                                   //current limit or reason for switch off output 6
                                   IF #statHMI.stateOutput6 = #CONST_STATE_OUT_AUTO_SWITCHED_OFF OR
                                       #statHMI.stateOutput6 = #CONST_STATE_OUT_RESET_POSSIBLE
                                   THEN
                                       #statHMI.reasonOutputSwitchedOff6 := BYTE_TO_INT(#statOutputCurrentLimit6);
                                   ELSE
                                       #statHMI.outputCurrentLimit6 := (BYTE_TO_INT(#statOutputCurrentLimit6) * #statHMI.nominalOutputCurrent) / #CONST_CONVERT_CURRENT;
                                   END_IF;

                                   //current limit or reason for switch off output 7
                                   IF #statHMI.stateOutput7 = #CONST_STATE_OUT_AUTO_SWITCHED_OFF OR
                                       #statHMI.stateOutput7 = #CONST_STATE_OUT_RESET_POSSIBLE
                                   THEN
                                       #statHMI.reasonOutputSwitchedOff7 := BYTE_TO_INT(#statOutputCurrentLimit7);
                                   ELSE
                                       #statHMI.outputCurrentLimit7 := (BYTE_TO_INT(#statOutputCurrentLimit7) * #statHMI.nominalOutputCurrent) / #CONST_CONVERT_CURRENT;
                                   END_IF;

                                   //current limit or reason for switch off output 8
                                   IF #statHMI.stateOutput8 = #CONST_STATE_OUT_AUTO_SWITCHED_OFF OR
                                       #statHMI.stateOutput8 = #CONST_STATE_OUT_RESET_POSSIBLE
                                   THEN
                                       #statHMI.reasonOutputSwitchedOff8 := BYTE_TO_INT(#statOutputCurrentLimit8);
                                   ELSE
                                       #statHMI.outputCurrentLimit8 := (BYTE_TO_INT(#statOutputCurrentLimit8) * #statHMI.nominalOutputCurrent) / #CONST_CONVERT_CURRENT;
                                   END_IF;

                               END_IF;

                           ELSE
                               // wrong frame Id
                               #statErrorFrameID := true;
                           END_IF;

                           IF #statGetFrame.frame0 = TRUE
                               AND #statGetFrame.frame1 = TRUE
                               AND #statGetFrame.frame2 = TRUE
                               AND #statGetFrame.frame3 = TRUE
                           THEN

                               #statIndexArticleNumber := 1;

                               FOR #statIndexArticleNumber := #CONST_START_CNT_INDEX1 TO #CONST_END_CNT_INDEX18 BY 1 DO
                                   IF #statArticleNumber[#statIndexArticleNumber] <> #statArticleNumberOld[#statIndexArticleNumber]
                                   THEN
                                       #statNewArticleNumberDetected := true;
                                   END_IF;
                               END_FOR;


                               IF #statNewArticleNumberDetected = TRUE
                               THEN

                                   #statNewArticleNumberDetected := false;
                                   #statArticleNumberChanged := true;

                                   Chars_TO_Strg(Chars := #statArticleNumber,
                                                 pChars := 0,
                                                 Cnt := 0,
                                                 Strg => #statHMI.articleNumber);
                                   #statArticleNumberOld := #statArticleNumber;
                               END_IF;


                               IF #statFabricationPlace = TRUE
                               THEN
                                   //fabrication place: Sibiu
                                   #statSerialNumber[1] := 'Y';
                                   #statSerialNumber[2] := 'S';
                                   #statSerialNumber[3] := 'U';
                                   #statSerialNumber[4] := '/';
                                   #statSerialNumber[5] := #statConstructionYearChar;
                                   #statSerialNumber[6] := #statConstructionMonthChar;
                                   #statSerialNumber[7] := ' ';
                                   #statSerialNumber[8] := ' ';
                                   #statSerialNumber[9] := ' ';
                                   #statSerialNumber[10] := ' ';
                                   #statSerialNumber[11] := ' ';
                                   #statSerialNumber[12] := ' ';
                                   #statSerialNumber[13] := ' ';
                               ELSE
                                   //fabrication place: Vienna
                                   #statSerialNumber[1] := 'Q';
                                   #statSerialNumber[2] := '6';
                                   #statSerialNumber[3] := '/';
                                   #statSerialNumber[4] := #statConstructionYearChar;
                                   #statSerialNumber[5] := #statConstructionMonthChar;
                                   #statSerialNumber[6] := ' ';
                                   #statSerialNumber[7] := ' ';
                                   #statSerialNumber[8] := ' ';
                                   #statSerialNumber[9] := ' ';
                                   #statSerialNumber[10] := ' ';
                                   #statSerialNumber[11] := ' ';
                                   #statSerialNumber[12] := ' ';
                                   #statSerialNumber[13] := ' ';

                               END_IF;

                               #statIndexSerialNumber := 1;

                               FOR #statIndexSerialNumber := #CONST_START_CNT_INDEX1 TO #CONST_END_CNT_INDEX13 BY 1 DO
                                   IF #statSerialNumber[#statIndexSerialNumber] <> #statSerialNumberOld[#statIndexSerialNumber]
                                   THEN
                                       #statNewSerialNumberDetected := true;
                                   END_IF;
                               END_FOR;

                               IF #statNewSerialNumberDetected = TRUE
                               THEN
                                   #statNewSerialNumberDetected := false;
                                   Chars_TO_Strg(Chars := #statSerialNumber,
                                                 pChars := 0,
                                                 Cnt := 0,
                                                 Strg => #statHMI.serialNumber);
                                   #statSerialNumberOld := #statSerialNumber;
                               END_IF;

                               #statGetFrame.frame0 := FALSE;
                               #statGetFrame.frame1 := FALSE;
                               #statGetFrame.frame2 := FALSE;
                               #statGetFrame.frame3 := FALSE;
                           END_IF;

                           // set output data structure
                           #HMI.deviceName := #statHMI.deviceName;
                           #HMI.stateCOM := true;
                           #HMI.stateDipSwitchTD1 := #statHMI.stateDipSwitchTD1;
                           #HMI.stateDipSwitchTD2 := #statHMI.stateDipSwitchTD2;
                           #HMI.stateOutput1 := #statHMI.stateOutput1;
                           #HMI.stateOutput2 := #statHMI.stateOutput2;
                           #HMI.stateOutput3 := #statHMI.stateOutput3;
                           #HMI.stateOutput4 := #statHMI.stateOutput4;
                           #HMI.stateOutput5 := #statHMI.stateOutput5;
                           #HMI.stateOutput6 := #statHMI.stateOutput6;
                           #HMI.stateOutput7 := #statHMI.stateOutput7;
                           #HMI.stateOutput8 := #statHMI.stateOutput8;
                           #HMI.outputCurrent1 := #statHMI.outputCurrent1;
                           #HMI.outputCurrent2 := #statHMI.outputCurrent2;
                           #HMI.outputCurrent3 := #statHMI.outputCurrent3;
                           #HMI.outputCurrent4 := #statHMI.outputCurrent4;
                           #HMI.outputCurrent5 := #statHMI.outputCurrent5;
                           #HMI.outputCurrent6 := #statHMI.outputCurrent6;
                           #HMI.outputCurrent7 := #statHMI.outputCurrent7;
                           #HMI.outputCurrent8 := #statHMI.outputCurrent8;
                           #HMI.outputCurrentLimit1 := #statHMI.outputCurrentLimit1;
                           #HMI.outputCurrentLimit2 := #statHMI.outputCurrentLimit2;
                           #HMI.outputCurrentLimit3 := #statHMI.outputCurrentLimit3;
                           #HMI.outputCurrentLimit4 := #statHMI.outputCurrentLimit4;
                           #HMI.outputCurrentLimit5 := #statHMI.outputCurrentLimit5;
                           #HMI.outputCurrentLimit6 := #statHMI.outputCurrentLimit6;
                           #HMI.outputCurrentLimit7 := #statHMI.outputCurrentLimit7;
                           #HMI.outputCurrentLimit8 := #statHMI.outputCurrentLimit8;
                           #HMI.reasonOutputSwitchedOff1 := #statHMI.reasonOutputSwitchedOff1;
                           #HMI.reasonOutputSwitchedOff2 := #statHMI.reasonOutputSwitchedOff2;
                           #HMI.reasonOutputSwitchedOff3 := #statHMI.reasonOutputSwitchedOff3;
                           #HMI.reasonOutputSwitchedOff4 := #statHMI.reasonOutputSwitchedOff4;
                           #HMI.reasonOutputSwitchedOff5 := #statHMI.reasonOutputSwitchedOff5;
                           #HMI.reasonOutputSwitchedOff6 := #statHMI.reasonOutputSwitchedOff6;
                           #HMI.reasonOutputSwitchedOff7 := #statHMI.reasonOutputSwitchedOff7;
                           #HMI.reasonOutputSwitchedOff8 := #statHMI.reasonOutputSwitchedOff8;
                           #HMI.nominalOutputCurrent := #statHMI.nominalOutputCurrent;
                           #HMI.productState := #statHMI.productState;
                           #HMI.firmwareVersion := #statHMI.firmwareVersion;
                           #HMI.startup := #statHMI.startup;
                           #HMI.outputNumber := #statHMI.outputNumber;
                           #HMI.stateReset := #statHMI.stateReset;
                           #HMI.articleNumber := #statHMI.articleNumber;
                           #HMI.serialNumber := #statHMI.serialNumber;

                       ELSE
                           //wrong device (no PSU OR SEL)
                           #statErrorDevice := true;
                       END_IF;
                       #statFrameOld := #statFrame;
                   END_IF;

               ELSE

                   IF #statInit = true
                   THEN
                       #statErrorFrameLength := true;
                   END_IF;

               END_IF;


               #statArrayImpulse[0] := #statTimeSave.deltaTimeImpulse;

               FOR #statIndexResetImpulse := #CONST_START_CNT_INDEX1 TO #CONST_END_CNT_INDEX63 BY 1 DO
                   #statArrayImpulse[#statIndexResetImpulse] := #CONST_TIME_0;
               END_FOR;

               FOR #statIndexResetPause := #CONST_START_CNT_INDEX0 TO #CONST_END_CNT_INDEX63 BY 1 DO
                   #statArrayPause[#statIndexResetPause] := #CONST_TIME_0;
               END_FOR;

               #statStartTimerWait := true;
               #statNoEvaluation := true;

               //Impulse detection    
           ELSIF #statTimeSave.deltaTimeImpulse >= #CONST_IMPULSE_MIN
               AND #statTimeSave.deltaTimeImpulse <= #CONST_IMPULSE_MAX
               AND #statImpulseDetected = TRUE
           THEN
               #statImpulseDetected := false;
               #statIndexResetImpulse := #CONST_INT_1;

               //save time of impulses to check frame length
               #statArrayImpulse[#statIndexImpulse] := #statTimeSave.deltaTimeImpulse;
               #statIndexImpulse := #statIndexImpulse + #CONST_INT_1;

               //count number of impulses
               #statCntImpulse := #statCntImpulse + #CONST_INT_1;

           END_IF;


           IF #statPauseDetected = TRUE
           THEN
               #statPauseDetected := false;
               #statIndexResetPause := #CONST_INT_0;

               //save time of pauses to check frame length
               #statArrayPause[#statIndexPause] := #statTimeSave.deltaTimePause;
               #statIndexPause := #statIndexPause + #CONST_INT_1;

               //count number of pauses
               #statCntPause := #statCntPause + #CONST_INT_1;

           END_IF;

           // bit detection
           IF #statNoEvaluation = false
               AND #statFrameEvaluationStopp = false
               AND ((#statPosEdgeDetectedTrigger = true)
               OR (#statNegEdgeDetectedTrigger = true))
           THEN

               IF #statPosEdgeDetectedTrigger = true
               THEN
                   #statArrayBits[#statCntBits] := true;
               ELSIF #statNegEdgeDetectedTrigger = true
               THEN
                   #statArrayBits[#statCntBits] := false;
               END_IF;

               #statStartTimerWait := true;
               #statNoEvaluation := true;

               IF (#statCntBits >= (#CONST_CNT_BITS_MAX - #CONST_INT_1))
               THEN
                   #statFrameEvaluationStopp := true;
                   #statCntBits := #CONST_INT_0;
               ELSE
                   #statCntBits := #statCntBits + #CONST_INT_1;
               END_IF;

           END_IF;

           //check max number of impulses and pauses in frame
           IF #statCntImpulse > #CONST_CNT_BITS_MAX
           THEN
               #statIndexImpulse := #CONST_INT_1;
               #statErrorFrameContent := TRUE;
           END_IF;

           IF #statCntPause > #CONST_CNT_PAUSE_MAX
           THEN
               #statIndexPause := #CONST_INT_0;
               #statErrorFrameContent := true;
           END_IF;

           IF #statErrorFrameContent = TRUE
           THEN
               #statStatusInt := #CONST_ERR_FRAMECONTENT;
               #statErrorInt := true;
           ELSIF #statErrorFrameLength = TRUE
           THEN
               #statStatusInt := #CONST_ERR_FRAMELENGTH;
               #statErrorInt := true;
           ELSIF #statErrorDevice = TRUE
           THEN
               #statStatusInt := #CONST_ERR_DEVICE;
               #statErrorInt := true;
           ELSIF #statErrorFrameID = TRUE
           THEN
               #statStatusInt := #CONST_ERR_FRAME_ID;
               #statErrorInt := true;
           ELSIF #statArticleNumberChanged = TRUE
           THEN
               #statStatusInt := #CONST_ERR_ARTICLE_NUMBER;
               #statErrorInt := true;
           END_IF;

           IF #statErrorInt = TRUE
           THEN
               #statErrorFrameLength := false;
               #statErrorFrameContent := false;
               #statErrorDevice := false;
               #statErrorFrameID := FALSE;
               #statArticleNumberChanged := false;
               #statStateIndex := #STATE_ERROR;
           END_IF;

       #STATE_ERROR:
           #statError := true;
           #statBusy := false;
           #statDone := false;
           #statStatus := #statStatusInt;
           #statStatusInt := #CONST_WORD_0;
           #statStartTimerSys := false;
           #statIndexResetBitArray := #CONST_INT_0;
           #statStartWatchDogTimerNeg := false;
           #statStartWatchDogTimerPos := false;

           IF #statErrorInt = TRUE
           THEN
               #statStateIndex := #STATE_EVALUATION;
               #statErrorInt := false;
               #statStartWatchDogTimerNeg := true;
               #statStartWatchDogTimerPos := true;
           ELSE
               #statStateIndex := #STATE_IDLE;
           END_IF;

       ELSE  // Statement section ELSE
           #statIndexResetBitArray := #CONST_INT_0;
           #statStateIndex := #STATE_IDLE;
   END_CASE;


   //Timer
   #instTimerWait(IN := #statStartTimerWait,
                  PT := #CONST_TIME_WAIT);

   IF #instTimerWait.Q = TRUE
   THEN
       #statStartTimerWait := false;
       #statNoEvaluation := false;
   END_IF;

   #instSysTimer(IN := #statStartTimerSys,
                 PT := #CONST_SYS_TIMER);


   IF #instSysTimer.Q = TRUE
   THEN
       #statStatusInt := #CONST_ERR_CYCLE_TIME;
       #statStateIndex := #STATE_ERROR;
   END_IF;

   #instWatchDogTimerPos(IN := #statStartWatchDogTimerPos,
                         PT := #CONST_WATCHDOG_TIMER);

   #instWatchDogTimerNeg(IN := #statStartWatchDogTimerNeg,
                         PT := #CONST_WATCHDOG_TIMER);

   IF #instWatchDogTimerNeg.Q = TRUE
       OR #instWatchDogTimerPos.Q = TRUE
   THEN
       #statStatusInt := #CONST_ERR_WATCHDOG;
       #statStateIndex := #STATE_ERROR;

       IF #HMI.stateNoCommunication = FALSE
       THEN
           #HMI.stateNoCommunication := true;

           #HMI.deviceName := #CONST_DEVICE_NAME_DEFAULT;
           #HMI.stateCOM := true;
           #HMI.stateDipSwitchTD1 := FALSE;
           #HMI.stateDipSwitchTD2 := FALSE;
           #HMI.stateOutput1 := #CONST_STATE_OUT_DEFAULT;
           #HMI.stateOutput2 := #CONST_STATE_OUT_DEFAULT;
           #HMI.stateOutput3 := #CONST_STATE_OUT_DEFAULT;
           #HMI.stateOutput4 := #CONST_STATE_OUT_DEFAULT;
           #HMI.stateOutput5 := #CONST_STATE_OUT_DEFAULT;
           #HMI.stateOutput6 := #CONST_STATE_OUT_DEFAULT;
           #HMI.stateOutput7 := #CONST_STATE_OUT_DEFAULT;
           #HMI.stateOutput8 := #CONST_STATE_OUT_DEFAULT;
           #HMI.outputCurrent1 := #CONST_CURRENT_OUT_DEFAULT;
           #HMI.outputCurrent2 := #CONST_CURRENT_OUT_DEFAULT;
           #HMI.outputCurrent3 := #CONST_CURRENT_OUT_DEFAULT;
           #HMI.outputCurrent4 := #CONST_CURRENT_OUT_DEFAULT;
           #HMI.outputCurrent5 := #CONST_CURRENT_OUT_DEFAULT;
           #HMI.outputCurrent6 := #CONST_CURRENT_OUT_DEFAULT;
           #HMI.outputCurrent7 := #CONST_CURRENT_OUT_DEFAULT;
           #HMI.outputCurrent8 := #CONST_CURRENT_OUT_DEFAULT;
           #HMI.outputCurrentLimit1 := #CONST_CURRENT_OUT_DEFAULT;
           #HMI.outputCurrentLimit2 := #CONST_CURRENT_OUT_DEFAULT;
           #HMI.outputCurrentLimit3 := #CONST_CURRENT_OUT_DEFAULT;
           #HMI.outputCurrentLimit4 := #CONST_CURRENT_OUT_DEFAULT;
           #HMI.outputCurrentLimit5 := #CONST_CURRENT_OUT_DEFAULT;
           #HMI.outputCurrentLimit6 := #CONST_CURRENT_OUT_DEFAULT;
           #HMI.outputCurrentLimit7 := #CONST_CURRENT_OUT_DEFAULT;
           #HMI.outputCurrentLimit8 := #CONST_CURRENT_OUT_DEFAULT;
           #HMI.reasonOutputSwitchedOff1 := #CONST_REASON_SWITCHED_OFF_DEFAULT;
           #HMI.reasonOutputSwitchedOff2 := #CONST_REASON_SWITCHED_OFF_DEFAULT;
           #HMI.reasonOutputSwitchedOff3 := #CONST_REASON_SWITCHED_OFF_DEFAULT;
           #HMI.reasonOutputSwitchedOff4 := #CONST_REASON_SWITCHED_OFF_DEFAULT;
           #HMI.reasonOutputSwitchedOff5 := #CONST_REASON_SWITCHED_OFF_DEFAULT;
           #HMI.reasonOutputSwitchedOff6 := #CONST_REASON_SWITCHED_OFF_DEFAULT;
           #HMI.reasonOutputSwitchedOff7 := #CONST_REASON_SWITCHED_OFF_DEFAULT;
           #HMI.reasonOutputSwitchedOff8 := #CONST_REASON_SWITCHED_OFF_DEFAULT;
           #HMI.nominalOutputCurrent := #CONST_NOMINAL_CURRENT3;
           #HMI.productState := #CONST_FW_PRODUCT_STATE_DEFAULT;
           #HMI.firmwareVersion := #CONST_FW_PRODUCT_STATE_DEFAULT;
           #HMI.startup := #CONST_STARTUP_DEFAULT;
           #HMI.outputNumber := #CONST_OUTPUT_NUMBER_4;
           #HMI.stateReset := FALSE;
           #HMI.articleNumber := #CONST_ARTICLE_NUMBER_DEFAULT;
           #HMI.serialNumber := #CONST_SERIAL_NUMBER_DEFAULT;

       END_IF;

   END_IF;

   #instTimerReset(IN:=#reset,
                   PT:=#CONST_RESET_TIMER);


   //edge Control
   #statImpulseOld := #impulse;
   #statPosEdgeDetectedTrigger := false;
   #statNegEdgeDetectedTrigger := false;

   //Cycle Time Control
   #statTimeSave.sysTimeOld := #statTimeSave.sysTime;

   // set outputs
   IF #HMI.setReset = TRUE
   THEN
       #HMI.setReset := false;
       #reset := true;
   ELSE
       IF #instTimerReset.Q = TRUE
       THEN
           #reset := false;
       END_IF;
   END_IF;

   #busy := #statBusy;
   #error := #statError;
   #done := #statDone;
   #status := #statStatus;
END_REGION
END_FUNCTION_BLOCK

FUNCTION_BLOCK "LPSE"   // FB6970, LAD
{ S7_Optimized_Access := 'TRUE' }
VERSION : 0.1
   VAR_INPUT
      impulse : Bool;
      reset : Bool;
   END_VAR
   VAR_OUTPUT
      done : Bool;
      busy : Bool;
      status : Word;
      error : Bool;
   END_VAR
   VAR
      statImpulseOld : Bool;
      HMI : Struct
         channelstate : Byte;
      END_STRUCT;
      statResetOld : Bool;
      statTimeSaver : Struct
         TimeTckRisingEdge : DTL;
         TimeTckFallingEdge : DTL;
         RisingEdgeDetected : Bool;
         FallingEdgeDetected : Bool;
         stateEdge : Int := 0;
      END_STRUCT;
      statDeltaTimeImpulse : Time;
      statDeltaTimePause : Time;
      statStartImpulseDetected : Bool;
      statImpulseDetected : Bool;
      statChannelState : Byte;
      statTimePauseSave0 : Time;
      statTimePauseSave1 : Time;
      statTimePauseSave2 : Time;
      statTimePauseSave3 : Time;
      statTimePauseSave4 : Time;
      statTimeImpulseSave0 : Time;
      statTimeImpulseSave1 : Time;
      statTimeImpulseSave2 : Time;
      statTimeImpulseSave3 : Time;
      statTimeImpulseSave4 : Time;
      statFrameImulseDetected : Bool;
      statNumberOfImpulses : Int;
      statChannelActive1 : Bool;
      statChannelActive2 : Bool;
      statChannelActive3 : Bool;
      statChannelActive4 : Bool;
      statCountChannelPos : Int;
      statCurrentPos1 : Int;
      statCurrentPos2 : Int;
      statCurrentPos3 : Int;
      statCurrentPos4 : Int;
      statTimeToImpulse : Time;
      statTimePause : Time;
      statTimeImpulse : Time;
      statTimeFrame : Time;
      statFrameOk : Bool;
      statCycleTimeNok : Bool;
      statDeltaSysTime : Time;
      instSysTimer : TON_TIME;
      statSysTimerStart : Bool;
      statSysTimerStop : Bool;
      statStatus : Word;
      statIndex : Int;
      statSysTimerRun : Time;
      instWatchDogTimerRising : TON_TIME;
      statWatchDogTimerRisingStart : Bool;
      statWatchDogTimerRisingStop : Bool;
      statWatchDogTimerRisingRun : Time;
      statResetRequest : Bool;
      statSysTimeDtl : DTL;
      statSysTimeOldDtl : DTL;
      instWatchDogTimerFalling : TON_TIME;
      statWatchDogTimerFallingStart : Bool;
      statWatchDogTimerFallingStop : Bool;
      statWatchDogTimerFallingRun : Time;
   END_VAR
   VAR_TEMP
      tempRetvalRdSys : Int;
      tempRetvalRdSysPosEdge : Int;
      tempRetvalRdSysNegEdge : Int;
      tempLatchTime : DTL;
      tempSysTime : DTL;
   END_VAR
   VAR CONSTANT
      STATE_IDLE : Int := 0;
      STATE_EVALUATION : Int := 1;
      STATE_ERROR : Int := 2;
      TIME_FRAME_MAX : Time := T#2850ms;
      TIME_FRAME_MIN : Time := T#2650ms;
      TIME_STARTIMPULSE_MIN : Time := T#400ms;
      TIME_STARTIMPULSE_MAX : Time := T#600ms;
      TIME_IMPULSE_MIN : Time := T#150ms;
      TIME_IMPULSE_MAX : Time := T#350ms;
      TIME_PAUSE1_MIN : Time := T#150ms;
      TIME_PAUSE1_MAX : Time := T#350ms;
      TIME_PAUSE2_MIN : Time := T#650ms;
      TIME_PAUSE2_MAX : Time := T#850ms;
      TIME_PAUSE3_MIN : Time := T#1150ms;
      TIME_PAUSE3_MAX : Time := T#1350ms;
      TIME_PAUSE4_MIN : Time := T#1650ms;
      TIME_PAUSE4_MAX : Time := T#1850ms;
      TIME_PAUSE_FRAME_MAX : Time := T#2350ms;
      TIME_PAUSE_FRAME_MIN : Time := T#2150ms;
      CONST_TIME_102 : Time := T#102ms;
      CONST_TIME_0 : Time := t#0ms;
      CONST_STATE_RISING_EDGE : Int := 15;
      CONST_STATE_FALLING_EDGE : Int := 16;
      CONST_WORD_0 : Word := 16#0000;
      CONST_BYTE_0 : Byte := 16#00;
      CONST_INT_0 : Int := 0;
      CONST_CHANNEL_POS4 : Int := 4;
      CONST_CHANNEL_POS1 : Int := 1;
      CONST_CHANNEL_POS2 : Int := 2;
      CONST_CHANNEL_POS3 : Int := 3;
      CONST_WATCHDOG_TIMER : Time := T#6s;
      CONST_CYCLETIME_TIMER : Time := T#4s;
      CONST_ERROR_CYCLETIME_TIMER : Word := 16#8001;
      CONST_ERROR_WATCHDOG_TIMER : Word := 16#8002;
   END_VAR
BEGIN

REGION Network 1 (SCL)
   //=============================================================================
   //SIEMENES AG
   //(c)Copyright 2017 All Rights Reserved
   //-----------------------------------------------------------------------------
   //Library:       LSitop
   //Tested with:   (S7-1200)
   //Engineering:    TIA Portal V15
   //Restrictions:   call in cyclic main OB
   //Requirements:
   //Functionality: evaluates the signal of status output (S) of SITOP PSE200U 
   //               ....
   //
   //-----------------------------------------------------------------------------
   //Change log table:
   //Version  Date       Expert in charge Changes applied
   //02.03.02 24.05.2017 (DI CS SD CSS KMT KD) Third released version
   //=============================================================================

   // Calculate cycle time

   // read date and time
   #tempRetvalRdSys := RD_SYS_T(#tempSysTime);
   #statSysTimeDtl := #tempSysTime;


   IF (#statSysTimeDtl > #statSysTimeOldDtl)
   THEN
       //calculate cycletime
       #statDeltaSysTime := T_DIFF(IN1 := #statSysTimeDtl, IN2 := #statSysTimeOldDtl);
       #statSysTimerStart := false;
   ELSE
       #statSysTimerStart := true;
       #statSysTimeOldDtl := #statSysTimeDtl;
       RETURN;
   END_IF;

   // check cycle time
   IF (#statDeltaSysTime >= #CONST_TIME_102)
   THEN
       #statCycleTimeNok := true;
       #statSysTimerStart := true;
   ELSE
       #statCycleTimeNok := false;
       #statSysTimerStart := false;
   END_IF;

   IF ((#reset = true)
       AND (#statResetOld = false))
   THEN
       #statSysTimerStart := false;
       #statWatchDogTimerRisingStart := false;
       #statWatchDogTimerFallingStart := false;
       #statResetRequest := true;
       #statIndex := #STATE_IDLE;
   END_IF;

   //Rising edge at impulse input
   IF ((#impulse = True)
       AND (#statImpulseOld = False))
   THEN
       #tempRetvalRdSysPosEdge := RD_SYS_T(#tempLatchTime);
       #statTimeSaver.RisingEdgeDetected := true;
       #statTimeSaver.stateEdge := #CONST_STATE_RISING_EDGE;
       #statTimeSaver.TimeTckRisingEdge := #tempLatchTime;
       #statWatchDogTimerRisingStart := true;
       #statWatchDogTimerFallingStart := false;

       IF (#busy = false)
       THEN
           #busy := true;
           #done := false;
           #error := false;
           #status := #CONST_WORD_0;
       END_IF;

       IF ((#statCycleTimeNok = false)
           AND (#statResetRequest = false))
       THEN
           #statIndex := #STATE_EVALUATION;
       END_IF;
   END_IF;

   //Falling edge at impulse input
   IF ((#impulse = False)
       AND (#statImpulseOld = True))
   THEN
       #tempRetvalRdSysNegEdge := RD_SYS_T(#tempLatchTime);
       #statTimeSaver.FallingEdgeDetected := true;
       #statTimeSaver.stateEdge := #CONST_STATE_FALLING_EDGE;
       #statTimeSaver.TimeTckFallingEdge := #tempLatchTime;
       #statWatchDogTimerFallingStart := true;
       #statWatchDogTimerRisingStart := false;

       IF ((#statCycleTimeNok = FALSE)
           AND (#statResetRequest = false))
       THEN
           #statIndex := #STATE_EVALUATION;
       END_IF;
   END_IF;

   IF ((#statTimeSaver.FallingEdgeDetected = false)
       AND (#statTimeSaver.RisingEdgeDetected = FALSE))
   THEN
       #statWatchDogTimerRisingStart := true;
       #statWatchDogTimerFallingStart := true;
   END_IF;

   CASE #statIndex OF
       #STATE_IDLE:  // IDLE_STATE
           #done := false;
           #error := false;
           #busy := false;
           #status := #CONST_WORD_0;
           #statStatus := #CONST_WORD_0;
           #HMI.channelstate := #CONST_BYTE_0;
           #statChannelState := #CONST_BYTE_0;
           #statFrameOk := false;
           #statCycleTimeNok := false;
           #statStartImpulseDetected := false;
           #statFrameImulseDetected := false;
           #statResetRequest := false;
           #statTimeSaver.FallingEdgeDetected := false;
           #statTimeSaver.RisingEdgeDetected := false;

       #STATE_EVALUATION:  //State: impulse detection

           //Delta time calculation
           IF ((#statTimeSaver.RisingEdgeDetected = True)
               AND (#statTimeSaver.FallingEdgeDetected = True))
           THEN

               IF (#statTimeSaver.stateEdge = #CONST_STATE_RISING_EDGE) //pos. edge, evaluate delta pause
               THEN

                   #statDeltaTimePause := T_DIFF(IN1 := #statTimeSaver.TimeTckRisingEdge, IN2 := #statTimeSaver.TimeTckFallingEdge);

                   IF ((#statDeltaTimePause < #CONST_TIME_0)
                       OR (#statDeltaTimePause > #TIME_FRAME_MAX))
                   THEN
                       #statIndex := #STATE_IDLE;
                       #statTimeSaver.FallingEdgeDetected := false;
                       RETURN;
                   END_IF;
                   #statTimeSaver.FallingEdgeDetected := false;

               END_IF;

               IF (#statTimeSaver.stateEdge = #CONST_STATE_FALLING_EDGE) // neg. edge, evaluate delta impulse
               THEN
                   #statImpulseDetected := true;
                   #statDeltaTimeImpulse := T_DIFF(IN1 := #statTimeSaver.TimeTckFallingEdge, IN2 := #statTimeSaver.TimeTckRisingEdge);

                   IF ((#statDeltaTimeImpulse < #CONST_TIME_0)
                       OR (#statDeltaTimeImpulse > #TIME_FRAME_MAX))
                   THEN
                       #statIndex := #STATE_IDLE;
                       #statTimeSaver.RisingEdgeDetected := false;
                       RETURN;
                   END_IF;
                   #statTimeSaver.RisingEdgeDetected := false;
               END_IF;

           END_IF;

           //Start bit detection
           IF ((#statDeltaTimeImpulse >= #TIME_STARTIMPULSE_MIN)
               AND (#statDeltaTimeImpulse <= #TIME_STARTIMPULSE_MAX))
               AND (#statImpulseDetected = True)
           THEN
               #statImpulseDetected := False;
               #statNumberOfImpulses := #CONST_INT_0;
               #statCountChannelPos := #CONST_INT_0;

               IF (#statCurrentPos1 = #CONST_INT_0)
               THEN
                   #statTimeImpulseSave1 := #CONST_TIME_0;
                   #statTimePauseSave1 := #CONST_TIME_0;
               END_IF;

               IF (#statCurrentPos2 = #CONST_INT_0)
               THEN
                   #statTimeImpulseSave2 := #CONST_TIME_0;
                   #statTimePauseSave2 := #CONST_TIME_0;
               END_IF;

               IF (#statCurrentPos3 = #CONST_INT_0)
               THEN
                   #statTimeImpulseSave3 := #CONST_TIME_0;
                   #statTimePauseSave3 := #CONST_TIME_0;
               END_IF;

               IF (#statCurrentPos4 = #CONST_INT_0)
               THEN
                   #statTimeImpulseSave4 := #CONST_TIME_0;
                   #statTimePauseSave4 := #CONST_TIME_0;
               END_IF;

               #statTimePauseSave0 := #statDeltaTimePause;
               #statTimeImpulseSave0 := #statDeltaTimeImpulse;

               // get time in sum of imulses
               #statTimeImpulse := #statTimeImpulseSave0 + #statTimeImpulseSave1 + #statTimeImpulseSave2 + #statTimeImpulseSave3 + #statTimeImpulseSave4;

               //get time in sum of pauses
               #statTimePause := #statTimePauseSave0 + #statTimePauseSave1 + #statTimePauseSave2 + #statTimePauseSave3 + #statTimePauseSave4;

               // get length of frame
               #statTimeFrame := #statTimeImpulse + #statTimePause;

               IF ((#statTimeFrame >= #TIME_FRAME_MIN)
                   AND (#statTimeFrame <= #TIME_FRAME_MAX)
                   AND (#statTimeToImpulse <= #TIME_FRAME_MAX))
               THEN
                   #statFrameOk := true;
               END_IF;

               IF ((#statFrameOk = TRUE)
                   AND (#statCycleTimeNok = FALSE))
               THEN
                   // Daten übernehmen
                   #done := true;
                   #busy := false;
                   #statFrameOk := false;

                   IF (#statChannelActive1 = true)
                   THEN
                       #statChannelState.%X0 := false;
                   ELSE
                       #statChannelState.%X0 := true;
                   END_IF;

                   IF (#statChannelActive2 = true)
                   THEN
                       #statChannelState.%X1 := false;
                   ELSE
                       #statChannelState.%X1 := true;
                   END_IF;

                   IF (#statChannelActive3 = true)
                   THEN
                       #statChannelState.%X2 := false;
                   ELSE
                       #statChannelState.%X2 := true;
                   END_IF;

                   IF (#statChannelActive4 = true)
                   THEN
                       #statChannelState.%X3 := false;
                   ELSE
                       #statChannelState.%X3 := true;
                   END_IF;

                   #HMI.channelstate := #statChannelState;
               END_IF;


               // channel 4 ok
               IF ((#statDeltaTimePause >= #TIME_PAUSE1_MIN)
                   AND (#statDeltaTimePause <= #TIME_PAUSE1_MAX))
               THEN
                   #statChannelActive4 := true;
                   // channel 4 ok not ok
               ELSIF ((#statDeltaTimePause >= #TIME_PAUSE2_MIN)
                   AND (#statDeltaTimePause <= #TIME_PAUSE2_MAX))
               THEN
                   #statChannelActive4 := false;
                   // channel 3 and 4 not ok    
               ELSIF ((#statDeltaTimePause >= #TIME_PAUSE3_MIN)
                   AND (#statDeltaTimePause <= #TIME_PAUSE3_MAX))
               THEN
                   #statChannelActive3 := false;
                   #statChannelActive4 := false;
                   // channel 2, 3, 4 not ok
               ELSIF ((#statDeltaTimePause >= #TIME_PAUSE4_MIN)
                   AND (#statDeltaTimePause <= #TIME_PAUSE4_MAX))
               THEN
                   #statChannelActive2 := false;
                   #statChannelActive3 := false;
                   #statChannelActive4 := false;
                   // channel 1, 2, 3, 4 not ok
               ELSIF ((#statDeltaTimePause >= #TIME_PAUSE_FRAME_MIN)
                   AND (#statDeltaTimePause <= #TIME_PAUSE_FRAME_MAX))
               THEN
                   #statChannelActive1 := false;
                   #statChannelActive2 := false;
                   #statChannelActive3 := false;
                   #statChannelActive4 := false;
               END_IF;

               #statCountChannelPos := #CONST_CHANNEL_POS4;

               #statCurrentPos1 := #CONST_INT_0;
               #statCurrentPos2 := #CONST_INT_0;
               #statCurrentPos3 := #CONST_INT_0;
               #statCurrentPos4 := #CONST_INT_0;

               // Imulse bit detection
           ELSIF ((#statDeltaTimeImpulse >= #TIME_IMPULSE_MIN)
               AND (#statDeltaTimeImpulse <= #TIME_IMPULSE_MAX))
               AND (#statImpulseDetected = True)
           THEN
               #statImpulseDetected := False;
               #statFrameImulseDetected := true;
           END_IF;

           //Channel detection

           IF (#statFrameImulseDetected = TRUE)
           THEN
               #statFrameImulseDetected := FALSE;

               IF (#statCountChannelPos = #CONST_CHANNEL_POS4)
               THEN
                   #statCurrentPos1 := #statCountChannelPos;
                   #statTimeImpulseSave1 := #statDeltaTimeImpulse;
                   #statTimePauseSave1 := #statDeltaTimePause;
                   #statTimeToImpulse := #CONST_TIME_0;
                   #statTimeToImpulse := #statTimeToImpulse + #statDeltaTimeImpulse + #statDeltaTimePause;

                   //channel 1 ok
                   IF ((#statDeltaTimePause >= #TIME_PAUSE1_MIN)
                       AND (#statDeltaTimePause <= #TIME_PAUSE1_MAX))
                   THEN
                       #statChannelActive1 := true;
                       #statCountChannelPos := #CONST_CHANNEL_POS1; // Pos 1 detected
                   END_IF;

                   // channel 1 not ok
                   IF ((#statDeltaTimePause >= #TIME_PAUSE2_MIN)
                       AND (#statDeltaTimePause <= #TIME_PAUSE2_MAX))
                   THEN
                       #statChannelActive1 := false;
                       #statChannelActive2 := true;
                       #statCountChannelPos := #CONST_CHANNEL_POS2; // go to next Pos 2
                   END_IF;

                   // channel 1 and 2 not ok
                   IF ((#statDeltaTimePause >= #TIME_PAUSE3_MIN)
                       AND (#statDeltaTimePause <= #TIME_PAUSE3_MAX))
                   THEN
                       #statChannelActive1 := false;
                       #statChannelActive2 := false;
                       #statChannelActive3 := true;
                       #statCountChannelPos := #CONST_CHANNEL_POS2; // go to next Pos 2
                   END_IF;

                   // channel 1, 2 and 3 not ok
                   IF ((#statDeltaTimePause >= #TIME_PAUSE4_MIN)
                       AND (#statDeltaTimePause <= #TIME_PAUSE4_MAX))
                   THEN
                       #statChannelActive1 := false;
                       #statChannelActive2 := false;
                       #statChannelActive3 := FALSE;
                       #statChannelActive4 := true;
                       #statCountChannelPos := #CONST_INT_0;
                   END_IF;

               ELSIF (#statCountChannelPos = #CONST_CHANNEL_POS1)
               THEN
                   #statCurrentPos2 := #statCountChannelPos;
                   #statTimeImpulseSave2 := #statDeltaTimeImpulse;
                   #statTimePauseSave2 := #statDeltaTimePause;
                   #statTimeToImpulse := #statTimeToImpulse + #statDeltaTimeImpulse + #statDeltaTimePause;

                   IF ((#statDeltaTimePause >= #TIME_PAUSE1_MIN)
                       AND (#statDeltaTimePause <= #TIME_PAUSE1_MAX))
                   THEN
                       #statChannelActive2 := true;
                       #statCountChannelPos := #CONST_CHANNEL_POS2; // go to next pos 2
                   END_IF;

                   IF ((#statDeltaTimePause >= #TIME_PAUSE2_MIN)
                       AND (#statDeltaTimePause <= #TIME_PAUSE2_MAX))
                   THEN
                       #statChannelActive2 := false;
                       #statChannelActive3 := true;
                       #statCountChannelPos := #CONST_CHANNEL_POS2; // go to next Pos 2
                   END_IF;

                   IF ((#statDeltaTimePause >= #TIME_PAUSE3_MIN)
                       AND (#statDeltaTimePause <= #TIME_PAUSE3_MAX))
                   THEN
                       #statChannelActive2 := false;
                       #statChannelActive3 := false;
                       #statChannelActive4 := true;
                       #statCountChannelPos := #CONST_INT_0;
                   END_IF;

               ELSIF (#statCountChannelPos = #CONST_CHANNEL_POS2)
               THEN
                   #statCurrentPos3 := #statCountChannelPos;
                   #statTimeImpulseSave3 := #statDeltaTimeImpulse;
                   #statTimePauseSave3 := #statDeltaTimePause;
                   #statTimeToImpulse := #statTimeToImpulse + #statDeltaTimeImpulse + #statDeltaTimePause;

                   IF ((#statDeltaTimePause >= #TIME_PAUSE1_MIN)
                       AND (#statDeltaTimePause <= #TIME_PAUSE1_MAX))
                   THEN
                       #statChannelActive3 := true;
                       #statCountChannelPos := #CONST_CHANNEL_POS3; // go to next pos 3
                   END_IF;

                   IF ((#statDeltaTimePause >= #TIME_PAUSE2_MIN)
                       AND (#statDeltaTimePause <= #TIME_PAUSE2_MAX))
                   THEN
                       #statChannelActive3 := false;
                       #statChannelActive4 := true;
                       #statCountChannelPos := #CONST_INT_0;
                   END_IF;

               ELSIF (#statCountChannelPos = #CONST_CHANNEL_POS3)
               THEN
                   #statCurrentPos4 := #statCountChannelPos;
                   #statTimeImpulseSave4 := #statDeltaTimeImpulse;
                   #statTimePauseSave4 := #statDeltaTimePause;
                   #statTimeToImpulse := #statTimeToImpulse + #statDeltaTimeImpulse + #statDeltaTimePause;

                   IF ((#statDeltaTimePause >= #TIME_PAUSE1_MIN)
                       AND (#statDeltaTimePause <= #TIME_PAUSE1_MAX))
                   THEN
                       #statChannelActive4 := true;
                   END_IF;
                   #statCountChannelPos := #CONST_INT_0; // go to pos 0
               END_IF;
           END_IF;

       #STATE_ERROR:
           #error := true;
           #busy := false;
           #done := false;
           #statSysTimerStart := false;
           #statWatchDogTimerRisingStart := false;
           #statWatchDogTimerFallingStart := false;
           #status := #statStatus;
           #statStatus := #CONST_WORD_0;
           #statIndex := #STATE_IDLE;
       ELSE
           #statIndex := #STATE_IDLE;
   END_CASE;

   #instWatchDogTimerRising(IN := #statWatchDogTimerRisingStart,
                            PT := #CONST_WATCHDOG_TIMER,
                            Q => #statWatchDogTimerRisingStop,
                            ET => #statWatchDogTimerRisingRun);


   #instWatchDogTimerFalling(IN:=#statWatchDogTimerFallingStart,
                             PT:=#CONST_WATCHDOG_TIMER,
                             Q=>#statWatchDogTimerFallingStop,
                             ET=>#statWatchDogTimerFallingRun);


   #instSysTimer(IN := #statSysTimerStart,
                 PT := #CONST_CYCLETIME_TIMER,
                 Q => #statSysTimerStop,
                 ET => #statSysTimerRun);

   IF (#statWatchDogTimerRisingStop = TRUE)
       OR (#statWatchDogTimerFallingStop = true)
   THEN
       #statIndex := #STATE_ERROR;
       #statStatus := #CONST_ERROR_WATCHDOG_TIMER;
   END_IF;


   IF (#statSysTimerStop = true)
   THEN
       #statIndex := #STATE_ERROR;
       #statStatus := #CONST_ERROR_CYCLETIME_TIMER;
   END_IF;

   //Edge control
   #statImpulseOld := #impulse;
   #statResetOld := #reset;

   // Cycle time control
   #statSysTimeOldDtl := #statSysTimeDtl;
END_REGION
END_FUNCTION_BLOCK

// folder: 1}Library/Simocode

FUNCTION_BLOCK "Simocode2"   // FB811, LAD
{ S7_Optimized_Access := 'TRUE' }